      CONST_RETAIN_TIME_SNAP_SIGNAL : Time := t#200ms;   // Time retain snap signal to z300
      CONST_DWRIDPLATE : DWord := 16#20002;   // R_ID message
      CONST_DWRIDMESSAGE2 : DWord := 16#30003;   // R_ID message
      CONST_DWRIDMESSAGE : DWord := 16#10001;   // R_ID message
      CONST_DGLASSBREAK_CLASS : DInt := 5;   // Glass break used class
      CONST_DGLASSBREAK_SUBTYPE : DInt := 1002;   // Glass break subtype
      CONST_DGLASSBREAK_DEFECT_WIDTH_CMM : DInt := 366000;   // Defect width [mm/100]
      CONST_DGLASSBREAK_DEFECT_GAP_CMM : DInt := 40000;   // Glass break defect gap [mm/100]
      CONST_DGLASSBREAK_LASTDEFECT_LENGTH_CMM : DInt := 50000;   // Last defect on glass break length [mm/100]
   END_VAR
BEGIN

REGION Network 1: ####_CONSTANTS_####
END_REGION

REGION Network 2: ####_MATCH_####
END_REGION

REGION Network 3 (SCL): General reset clean
   IF #IN_xGeneralReset THEN

       #TMP_dwValue := 0;

       SCATTER(IN:=#TMP_dwValue,
               OUT=>#tPhases);

       SCATTER(IN:=#TMP_dwValue,
               OUT=>#tPhasesNetworkPlate);


   END_IF;
END_REGION

REGION Network 4 (SCL): Move data information to tracking
   #INO_tTrack.rgtTrackMachine[#IN_dMachineIndex].tUserData.dSetDistanceSnap_cmm := #IN_dSnapOffset_cmm*-1;
   #INO_tTrack.rgtTrackMachine[#IN_dMachineIndex].tUserData.dSetMachReacTime_ms := #tHMW.dAccelerationDelay_ms;
END_REGION

REGION Network 5 (SCL): Manage tracking call

   #OS_xNewCapUp := FALSE;
   #OS_xNewCapDw := FALSE;
   #OS_xNewCap := FALSE;
   #OS_xNewCapFastDropUp := FALSE;
   IF #INO_tTrack.rgtTrackMachine[#IN_dMachineIndex].tUserData.xGetPosReach THEN

       IF (NOT #ST_xPhaseInProgress) THEN

           IF #INO_tTrack.rgtTrackMachine[#IN_dMachineIndex].tUserData.dGetUpstremIndex >= 0 THEN
               #AUX_dUpCapIndex := #INO_tTrack.rgtTrackMachine[#IN_dMachineIndex].tUserData.dGetUpstremIndex;
               IF #INO_tTrack.rgtTrackCaps[#AUX_dUpCapIndex].tCap.dLength_cmm >= #CONST_MINPLATELENGTH_Z300_CMM THEN
                   #OS_xNewCapUp := TRUE;
                   #AUX_xValidUpCap := TRUE;
               ELSE
                   #AUX_xValidUpCap := FALSE;

               END_IF;
           ELSE
                   #AUX_xValidUpCap := FALSE;
                   #OS_xNewCapUp := FALSE;
                   #AUX_dUpCapIndex := 0;
           END_IF;

           IF #INO_tTrack.rgtTrackMachine[#IN_dMachineIndex].tUserData.dGetDownstreamIndex >= 0 THEN
               #AUX_xValidDwCap := TRUE;
               #OS_xNewCapDw := TRUE;            
               #AUX_dDwCapIndex := #INO_tTrack.rgtTrackMachine[#IN_dMachineIndex].tUserData.dGetDownstreamIndex;

               IF #INO_tTrack.rgtTrackCaps[#AUX_dDwCapIndex].tCap.dLength_cmm >= #CONST_MINPLATELENGTH_Z300_CMM THEN
                   #OS_xNewCap := TRUE;
               ELSE
                   #OS_xNewCapFastDropUp := TRUE;
               END_IF;

           ELSE
               #AUX_xValidDwCap := FALSE;
               #OS_xNewCapDw := FALSE;            
               #AUX_dDwCapIndex := 0;
           END_IF;



       END_IF;

       #INO_tTrack.rgtTrackMachine[#IN_dMachineIndex].tUserData.xGetPosReach := FALSE;

   END_IF;
END_REGION

REGION Network 6 (SCL): Manage message
   IF #AUX_xValidUpCap AND (#OS_xNewCapUp OR  #OS_xNewCapFastDropUp) THEN

       //Evaluate the missing xcut, send to cullet the upstream and downstream. On the downstream send also the message
       #TMP_xCutDone := FALSE;
       #AUX_xXcutDone := FALSE;
       FOR #TMP_dIndex := 0 TO "DMAXXHEADS_IND" DO
           IF #INO_tTrack.rgtTrackCaps[#AUX_dUpCapIndex].tCap.tDone.rgxXCutDoneHead[#TMP_dIndex] THEN
               #TMP_xCutDone := TRUE;
               #AUX_xXcutDone := TRUE;
               EXIT;                    
           END_IF;
       END_FOR;

       IF #TMP_xCutDone = FALSE THEN  

           //Send to cullet the upstream
           FOR #TMP_dIndex := 0 TO  #INO_tTrack.rgtTrackCaps[#AUX_dUpCapIndex].tCap.dNumLites - 1 DO

               IF #INO_tTrack.rgtTrackCaps[#AUX_dUpCapIndex].tCap.rgtLites[#TMP_dIndex].dMainDestination <> "DCULLETDESTMASK" THEN

                   #INO_tTrack.rgtTrackCaps[#AUX_dUpCapIndex].tCap.rgtLites[#TMP_dIndex].dMainDestination := "DCULLETDESTMASK";
                   #INO_tTrack.rgtTrackCaps[#AUX_dUpCapIndex].tCap.rgtLites[#TMP_dIndex].dAltDestination := 0;
                   #INO_tTrack.rgtTrackCaps[#AUX_dUpCapIndex].tCap.rgtLites[#TMP_dIndex].d2ndDestionation := 0;
                   #INO_tTrack.rgtTrackCaps[#AUX_dUpCapIndex].tCap.rgtLites[#TMP_dIndex].dCulletCause := "DCULLETCAUSE_XCUTMISSING";

               END_IF;
           END_FOR;

           #INO_tTrack.rgtTrackCaps[#AUX_dUpCapIndex].tCap.tRequests.xUpdateDataBPSA := TRUE;
           #INO_tTrack.rgtTrackCaps[#AUX_dUpCapIndex].tCap.tRequests.xUpdateDataBPSB := TRUE;

           //Send to cullet the downstream
           FOR #TMP_dIndex := 0 TO  #INO_tTrack.rgtTrackCaps[#AUX_dDwCapIndex].tCap.dNumLites - 1 DO

               IF #INO_tTrack.rgtTrackCaps[#AUX_dDwCapIndex].tCap.rgtLites[#TMP_dIndex].dMainDestination <> "DCULLETDESTMASK" THEN

                   #INO_tTrack.rgtTrackCaps[#AUX_dDwCapIndex].tCap.rgtLites[#TMP_dIndex].dMainDestination := "DCULLETDESTMASK";
                   #INO_tTrack.rgtTrackCaps[#AUX_dDwCapIndex].tCap.rgtLites[#TMP_dIndex].dAltDestination := 0;
                   #INO_tTrack.rgtTrackCaps[#AUX_dDwCapIndex].tCap.rgtLites[#TMP_dIndex].d2ndDestionation := 0;
                   #INO_tTrack.rgtTrackCaps[#AUX_dDwCapIndex].tCap.rgtLites[#TMP_dIndex].dCulletCause := "DCULLETCAUSE_XCUTMISSING";

                   "RP_AddMessageV2"(IN_xInit:=FALSE,
                     IN_dCodeEvent:="DEVENTS_REDESTINATION",
                     IN_strIndet_Max4Chars:='Z200',
                     IN_dValue1:="DEVENTS_CULLETDESTINATION",
                     IN_dValue2:=#INO_tTrack.rgtTrackCaps[#AUX_dDwCapIndex].tCap.rgtLites[#TMP_dIndex].dID,
                     IN_dValue3:=#INO_tTrack.rgtTrackCaps[#AUX_dDwCapIndex].tCap.rgtLites[#TMP_dIndex].dProductionID,
                     IN_dValue4:=#INO_tTrack.rgtTrackCaps[#AUX_dDwCapIndex].tCap.rgtLites[#TMP_dIndex].dCulletCause,
                     IN_dValue5:=0,
                     IN_dValue6:=0,
                     IN_dValue7:=0,
                     IN_dValue8:=0,
                     IN_dValue9:=0,
                     IN_dValue10:=0,
                     INO_tBuffer:=#INO_tMessage,
                     INO_xError:=#INO_xMessageAnomaly);

               END_IF;
           END_FOR;

           #INO_tTrack.rgtTrackCaps[#AUX_dUpCapIndex].tCap.tRequests.xUpdateDataBPSA := TRUE;
           #INO_tTrack.rgtTrackCaps[#AUX_dUpCapIndex].tCap.tRequests.xUpdateDataBPSB := TRUE;

       END_IF;

       FOR #TMP_dIndex := 0 TO #INO_tTrack.rgtTrackCaps[#AUX_dUpCapIndex].tCap.dNumLites - 1 DO

           IF #INO_tTrack.rgtTrackCaps[#AUX_dUpCapIndex].tCap.rgtLites[#TMP_dIndex].dMainDestination = "DCULLETDESTMASK" THEN
              "RP_AddMessageV2"(IN_xInit:=FALSE,
                     IN_dCodeEvent:="DEVENTS_REDESTINATION",
                     IN_strIndet_Max4Chars:='Z200',
                     IN_dValue1:="DEVENTS_CULLETDESTINATION",
                     IN_dValue2:=#INO_tTrack.rgtTrackCaps[#AUX_dUpCapIndex].tCap.rgtLites[#TMP_dIndex].dID,
                     IN_dValue3:=#INO_tTrack.rgtTrackCaps[#AUX_dUpCapIndex].tCap.rgtLites[#TMP_dIndex].dProductionID,
                     IN_dValue4:=#INO_tTrack.rgtTrackCaps[#AUX_dUpCapIndex].tCap.rgtLites[#TMP_dIndex].dCulletCause,
                     IN_dValue5:=0,
                     IN_dValue6:=0,
                     IN_dValue7:=0,
                     IN_dValue8:=0,
                     IN_dValue9:=0,
                     IN_dValue10:=0,
                     INO_tBuffer:=#INO_tMessage,
                     INO_xError:=#INO_xMessageAnomaly);
           END_IF;


       END_FOR;

   END_IF;
END_REGION

REGION Network 7: ####_HMI_LOGICS_####
END_REGION

REGION Network 8 (SCL): List of HMI logics
END_REGION

REGION Network 9: ####_ALARMS_####
END_REGION

REGION Network 10 (SCL): Reset alarms
   IF #IN_xResetAlarms THEN

       #TMP_dwValue := 0;

       SCATTER(IN:=#TMP_dwValue,
               OUT=>#tALM.tF);

       SCATTER(IN:=#TMP_dwValue,
               OUT=>#tALM.tS);

       SCATTER(IN:=#TMP_dwValue,
               OUT=>#tALM.tW);

   END_IF;
END_REGION

REGION Network 11: ####_STATUSES_####
END_REGION

REGION Network 12 (SCL): Calculate alarm statuses
   GATHER(IN:=#tALM.tS,
          OUT=>#TMP_dwValue);

   IF #TMP_dwValue <> 0 THEN
       #ST_xStoppingFaults := TRUE;
   ELSE
       #ST_xStoppingFaults := FALSE;
   END_IF;

   GATHER(IN:=#tALM.tF,
          OUT=>#TMP_dwValue);

   IF #TMP_dwValue <> 0 THEN
       #ST_xFaults := TRUE;
   ELSE
       #ST_xFaults := FALSE;
   END_IF;

   GATHER(IN:=#tALM.tW,
          OUT=>#TMP_dwValue);

   IF #TMP_dwValue <> 0 THEN
       #ST_xWarnings := TRUE;
   ELSE
       #ST_xWarnings := FALSE;
   END_IF;
END_REGION

REGION Network 13: Send data request
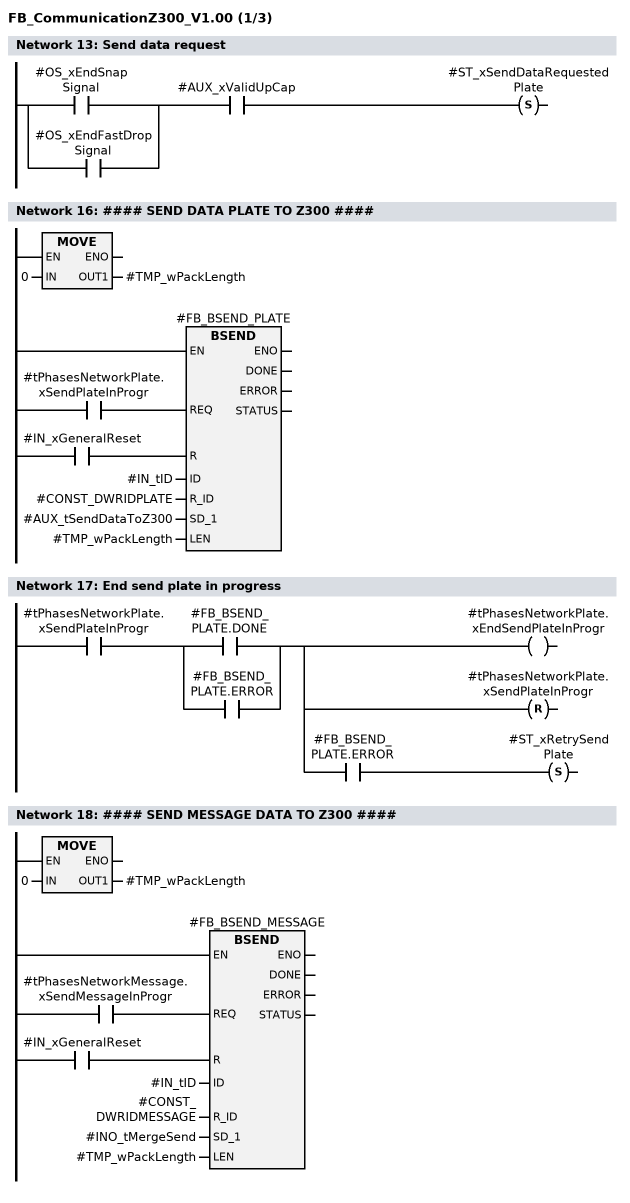
   RUNG wire#powerrail
      Contact( #OS_xEndSnapSignal )
      wire#w1
      Contact( #AUX_xValidUpCap )
      S_Coil( #ST_xSendDataRequestedPlate )
   END_RUNG
   RUNG wire#powerrail
      Contact( #OS_xEndFastDropSignal )
   END_RUNG wire#w1
   // the same network as SCL:
   IF (#OS_xEndSnapSignal OR #OS_xEndFastDropSignal) AND #AUX_xValidUpCap THEN
       #ST_xSendDataRequestedPlate := TRUE;
   END_IF;
END_REGION

REGION Network 14 (SCL): Compile Data for Z300
   IF NOT #ST_xPhaseInProgressNetworkPlate AND (#ST_xSendDataRequestedPlate OR #ST_xRetrySendPlate) THEN


       IF #ST_xSendDataRequestedPlate THEN

           //clean buffer
           #AUX_tSendDataToZ300 := #AUX_tEmptySendDataToZ300;
           //Convoy data.Search plate
           IF #INO_tTrack.rgtTrackCaps[#AUX_dUpCapIndex].tCap.dIndex = 0 THEN

               //Search until the previous cap
               #TMP_dIndex := 1;
               #TMP_dValue := #AUX_dUpCapIndex;
               #TMP_dConvNumPlate := 1;
               #TMP_dConvTotalLength_cmm := #INO_tTrack.rgtTrackCaps[#AUX_dUpCapIndex].tCap.dLength_cmm;

               WHILE #TMP_dIndex < "DMAXCAP_Z300" DO

                   #TMP_dValue := #TMP_dValue + 1;

                   IF #TMP_dValue > "DMAXTRACKCAP_IND" THEN
                       #TMP_dValue := 0;
                   END_IF;

                   IF #INO_tTrack.rgtTrackCaps[#TMP_dValue].tCap.dIndex <> 0 THEN

                       #TMP_dConvNumPlate := #TMP_dConvNumPlate + 1;
                       #TMP_dConvTotalLength_cmm := #TMP_dConvTotalLength_cmm + #INO_tTrack.rgtTrackCaps[#TMP_dValue].tCap.dLength_cmm;
                   ELSE

                       EXIT;

                   END_IF;

                   #TMP_dIndex := #TMP_dIndex + 1;

               END_WHILE;

               IF #TMP_dConvNumPlate > 1 THEN

                   //Convoy present, calculate gap.
                   #TMP_dConvGap_cmm := ("DMAXLENGHTCONVOY_CMM" - #TMP_dConvTotalLength_cmm) / (#TMP_dConvNumPlate - 1);
                   #TMP_dValue := #AUX_dUpCapIndex;
                   #TMP_dIndex := 0;
                   //Update plate data
                   WHILE (#TMP_dIndex < #TMP_dConvNumPlate) DO

                       #INO_tTrack.rgtTrackCaps[#TMP_dValue].tCap.dIndex := #TMP_dIndex;

                       IF (#TMP_dIndex + 1) < #TMP_dConvNumPlate THEN
                           #INO_tTrack.rgtTrackCaps[#TMP_dValue].tCap.dReqGapForConv_cmm := 50000; //#TMP_dConvGap_cmm;
                       ELSE
                           #INO_tTrack.rgtTrackCaps[#TMP_dValue].tCap.dReqGapForConv_cmm := 0;
                       END_IF;

                       #TMP_dIndex := #TMP_dIndex + 1;

                       #TMP_dValue := #TMP_dValue + 1;

                       IF #TMP_dValue > "DMAXTRACKCAP_IND"  THEN
                           #TMP_dValue := 0;
                       END_IF;

                   END_WHILE;
               END_IF;
           END_IF;

           #AUX_tCapToSend := #INO_tTrack.rgtTrackCaps[#AUX_dUpCapIndex].tCap;
           //compile plate data TO Z300
           #AUX_tSendDataToZ300.dID := #INO_tTrack.rgtTrackCaps[#AUX_dUpCapIndex].tCap.dID;
           #AUX_tSendDataToZ300.dProductionID := 1;
           #AUX_tSendDataToZ300.dLength_cmm := #INO_tTrack.rgtTrackCaps[#AUX_dUpCapIndex].tCap.dLength_cmm;
           #AUX_tSendDataToZ300.dWidth_cmm := #INO_tTrack.rgtTrackCaps[#AUX_dUpCapIndex].tCap.dWidth_cmm;
           #AUX_tSendDataToZ300.dThick_cmm := #INO_tTrack.rgtTrackCaps[#AUX_dUpCapIndex].tCap.dThick_cmm;
           #AUX_tSendDataToZ300.dIndex := #INO_tTrack.rgtTrackCaps[#AUX_dUpCapIndex].tCap.dIndex;
           #AUX_tSendDataToZ300.dFormat := #INO_tTrack.rgtTrackCaps[#AUX_dUpCapIndex].tCap.dFormat;
           #AUX_tSendDataToZ300.dNumLites := #INO_tTrack.rgtTrackCaps[#AUX_dUpCapIndex].tCap.dNumLites;

           #AUX_tSendDataToZ300.dReqGapForConv_cmm := 0;
           IF #INO_tTrack.rgtTrackCaps[#AUX_dUpCapIndex].tCap.dMaxCapInConv>1
               AND (#INO_tTrack.rgtTrackCaps[#AUX_dUpCapIndex].tCap.dMaxCapInConv-1>#AUX_tSendDataToZ300.dIndex) THEN
               #AUX_tSendDataToZ300.dReqGapForConv_cmm := 50000;
               #AUX_tSendDataToZ300.dGap_cmm := 50000;
           END_IF;
           #AUX_tSendDataToZ300.dMaxCapInConv := #INO_tTrack.rgtTrackCaps[#AUX_dUpCapIndex].tCap.dMaxCapInConv;

           #TMP_dValue := #AUX_dUpCapIndex + 1;

           IF #TMP_dValue >= "DMAXTRACKCAP_IND" THEN
               #TMP_dValue := 0;
           END_IF;
           IF #INO_tTrack.rgtTrackCaps[#TMP_dValue].tCap.dMaxCapInConv = 0 THEN
               #AUX_tSendDataToZ300.dReqGapForConv_cmm := 0;
               #AUX_tSendDataToZ300.dGap_cmm := 0;
               #AUX_tSendDataToZ300.dMaxCapInConv := 0;
           END_IF;


           #AUX_tSendDataToZ300.dConvTotLength_cmm := #INO_tTrack.rgtTrackCaps[#AUX_dUpCapIndex].tCap.dConvTotLength_cmm;
           #AUX_tSendDataToZ300.dMinWidth_cmm := #INO_tTrack.rgtTrackCaps[#AUX_dUpCapIndex].tCap.dMinWidth_cmm;
           #AUX_tSendDataToZ300.dMaxWidth_cmm := #INO_tTrack.rgtTrackCaps[#AUX_dUpCapIndex].tCap.dMaxWidth_cmm;
           #AUX_tSendDataToZ300.dGrossWidth_cmm := #INO_tTrack.rgtTrackCaps[#AUX_dUpCapIndex].tCap.dGrossWidth_cmm;
           #AUX_tSendDataToZ300.dNetWidth_cmm := #INO_tTrack.rgtTrackCaps[#AUX_dUpCapIndex].tCap.dNetWidth_cmm;
           #AUX_tSendDataToZ300.dDEdgeOpSide_cmm := #INO_tTrack.rgtTrackCaps[#AUX_dUpCapIndex].tCap.dDEdgeOpSide_cmm;
           #AUX_tSendDataToZ300.dDEdgeOppOpSide_cmm := #INO_tTrack.rgtTrackCaps[#AUX_dUpCapIndex].tCap.dDEdgeOppOpSide_cmm;
           #AUX_tSendDataToZ300.dTEdgeOpSide_cmm := #INO_tTrack.rgtTrackCaps[#AUX_dUpCapIndex].tCap.dTEdgeOpSide_cmm;
           #AUX_tSendDataToZ300.dTEdgeOppOpSide_cmm := #INO_tTrack.rgtTrackCaps[#AUX_dUpCapIndex].tCap.dTEdgeOppOpSide_cmm;
           #AUX_tSendDataToZ300.dCutWander_cmm := #INO_tTrack.rgtTrackCaps[#AUX_dUpCapIndex].tCap.dEndCutWander_cmm;
           #AUX_tSendDataToZ300.dColor := #INO_tTrack.rgtTrackCaps[#AUX_dUpCapIndex].tCap.dColor;
           #AUX_tSendDataToZ300.strColorDescr := #INO_tTrack.rgtTrackCaps[#AUX_dUpCapIndex].tCap.strColorDescr;

           #TMP_xReqDoneMatch := FALSE;
           GATHER(IN :=  #INO_tTrack.rgtTrackCaps[#AUX_dUpCapIndex].tCap.tDone.tYCuts[0].rgxHeadsDone,
                  OUT => #TMP_wValue);
           IF #TMP_wValue <> 0 THEN
               #AUX_tSendDataToZ300.tFlagTrim.xByYCut1 := TRUE;

               IF #INO_tTrack.rgtTrackCaps[#AUX_dUpCapIndex].tCap.tDone.tYCuts[0].rgxHeadsDone = 
                       #INO_tTrack.rgtTrackCaps[#AUX_dUpCapIndex].tCap.tRequests.tYCutsData[0].rgxHeadsRequest THEN
                   #TMP_xReqDoneMatch := TRUE;
               END_IF;

           END_IF;
           GATHER(IN := #INO_tTrack.rgtTrackCaps[#AUX_dUpCapIndex].tCap.tDone.tYCuts[1].rgxHeadsDone,
                  OUT => #TMP_wValue);
           IF #TMP_wValue <> 0 THEN
               #AUX_tSendDataToZ300.tFlagTrim.xByYCut2 := TRUE;

               IF #INO_tTrack.rgtTrackCaps[#AUX_dUpCapIndex].tCap.tDone.tYCuts[1].rgxHeadsDone = 
                       #INO_tTrack.rgtTrackCaps[#AUX_dUpCapIndex].tCap.tRequests.tYCutsData[1].rgxHeadsRequest THEN
                   #TMP_xReqDoneMatch := TRUE;
               END_IF;

           END_IF;

           IF #TMP_xReqDoneMatch THEN

               IF #INO_tTrack.rgtTrackCaps[#AUX_dUpCapIndex].tCap.dTEdgeOpSide_cmm > 0 THEN
                   #AUX_tSendDataToZ300.tFlagTrim.xTrim3OpSide := 1;
               END_IF;
               IF #INO_tTrack.rgtTrackCaps[#AUX_dUpCapIndex].tCap.dDEdgeOpSide_cmm > 0 THEN
                   #AUX_tSendDataToZ300.tFlagTrim.xTrim2OpSide := 1;
               END_IF;

               #AUX_tSendDataToZ300.tFlagTrim.xTrim1OpSide := 1;
               #AUX_tSendDataToZ300.tFlagTrim.xTrim1OppOpSide := 1;

               IF #INO_tTrack.rgtTrackCaps[#AUX_dUpCapIndex].tCap.dDEdgeOppOpSide_cmm > 0 THEN
                   #AUX_tSendDataToZ300.tFlagTrim.xTrim2OppOpSide := 1;
               END_IF;
               IF #INO_tTrack.rgtTrackCaps[#AUX_dUpCapIndex].tCap.dTEdgeOppOpSide_cmm > 0 THEN
                   #AUX_tSendDataToZ300.tFlagTrim.xTrim3OppOpSide := 1;
               END_IF;

               FOR #TMP_dIndex := 1 TO #INO_tTrack.rgtTrackCaps[#AUX_dUpCapIndex].tCap.dNumLites - 1 DO
                   #AUX_tSendDataToZ300.tFlagTrim.rgxIntCut[#TMP_dIndex - 1] := 1;
               END_FOR;

           ELSE
               #AUX_tSendDataToZ300.tFlagTrim.xTrim3OpSide := 0;
               #AUX_tSendDataToZ300.tFlagTrim.xTrim2OpSide := 0;
               #AUX_tSendDataToZ300.tFlagTrim.xTrim1OpSide := 0;
               #AUX_tSendDataToZ300.tFlagTrim.xTrim1OppOpSide := 0;
               #AUX_tSendDataToZ300.tFlagTrim.xTrim2OppOpSide := 0;
               #AUX_tSendDataToZ300.tFlagTrim.xTrim3OppOpSide := 0;
           END_IF;

           #AUX_tSendDataToZ300.tFlagTrim.xOptSelvedgeSel := #INO_tTrack.rgtTrackCaps[#AUX_dUpCapIndex].tCap.tRequests.xOptSelvedgeSel;
           #AUX_tSendDataToZ300.tFlagTrim.xOptSplitBarSel := #INO_tTrack.rgtTrackCaps[#AUX_dUpCapIndex].tCap.tRequests.xOptSplitBarSel;
           #AUX_tSendDataToZ300.tFlagTrim.xOptSepRollSel := #INO_tTrack.rgtTrackCaps[#AUX_dUpCapIndex].tCap.tRequests.xOptSepRollSel;

           FOR #TMP_dIndex := 0 TO "DMAXXHEADS_IND" DO
               #AUX_tSendDataToZ300.tFlagTrim.rgxXCutDoneHead[#TMP_dIndex] := #INO_tTrack.rgtTrackCaps[#AUX_dUpCapIndex].tCap.tDone.rgxXCutDoneHead[#TMP_dIndex];
           END_FOR;

           FOR #TMP_dIndex := 0 TO "DMAXXHEADS_IND" DO
               #AUX_tSendDataToZ300.tFlagTrim.rgxXCutDoneTail[#TMP_dIndex] := #INO_tTrack.rgtTrackCaps[#AUX_dUpCapIndex].tCap.tDone.rgxXCutDoneTail[#TMP_dIndex];
           END_FOR;

           IF #AUX_tSendDataToZ300.tFlagTrim.xByYCut1 THEN
               #AUX_tSendDataToZ300.tFlagTrim.rgxYCutHeadDone := #INO_tTrack.rgtTrackCaps[#AUX_dUpCapIndex].tCap.tDone.tYCuts[0].rgxHeadsDone;
           ELSE
               #AUX_tSendDataToZ300.tFlagTrim.rgxYCutHeadDone := #INO_tTrack.rgtTrackCaps[#AUX_dUpCapIndex].tCap.tDone.tYCuts[1].rgxHeadsDone;
           END_IF;

           #AUX_tSendDataToZ300.tFlagTrim.tSelvedge.dRequestTrim3OpSide := #INO_tTrack.rgtTrackCaps[#AUX_dUpCapIndex].tCap.tRequests.dReqTrim3OpSide;
           #AUX_tSendDataToZ300.tFlagTrim.tSelvedge.dRequestTrim2OpSide := #INO_tTrack.rgtTrackCaps[#AUX_dUpCapIndex].tCap.tRequests.dReqTrim2OpSide;
           #AUX_tSendDataToZ300.tFlagTrim.tSelvedge.dRequestTrim1OpSide := #INO_tTrack.rgtTrackCaps[#AUX_dUpCapIndex].tCap.tRequests.dReqTrim1OpSide;
           #AUX_tSendDataToZ300.tFlagTrim.tSelvedge.dRequestTrim3OppOpSide := #INO_tTrack.rgtTrackCaps[#AUX_dUpCapIndex].tCap.tRequests.dReqTrim3OppOpSide;
           #AUX_tSendDataToZ300.tFlagTrim.tSelvedge.dRequestTrim2OppOpSide := #INO_tTrack.rgtTrackCaps[#AUX_dUpCapIndex].tCap.tRequests.dReqTrim2OppOpSide;
           #AUX_tSendDataToZ300.tFlagTrim.tSelvedge.dRequestTrim1OppOpSide := #INO_tTrack.rgtTrackCaps[#AUX_dUpCapIndex].tCap.tRequests.dReqTrim1OppOpSide;

           FOR #TMP_dIndex := 0 TO "DMAXLITE_IND" DO
               #AUX_tSendDataToZ300.tFlagTrim.tSplitBar[#TMP_dIndex].dRequestSnapCut := #INO_tTrack.rgtTrackCaps[#AUX_dUpCapIndex].tCap.tRequests.rgdReqSplitBarSel[#TMP_dIndex];
           END_FOR;

           FOR #TMP_dIndex := 0 TO "DMAXSEPROLLBANK_IND" DO
               #TMP_wValue := INT_TO_WORD(#INO_tTrack.rgtTrackCaps[#AUX_dUpCapIndex].tCap.tRequests.rgbSeparatorSelect[#TMP_dIndex]);
               SCATTER(IN := #TMP_wValue,
                       OUT => #TMP_rgxWValue);
               #AUX_tSendDataToZ300.tFlagTrim.tSepRoll[#TMP_dIndex].rgxRequestSeparator := #TMP_rgxWValue;
           END_FOR;

           FOR #TMP_dIndex := 0 TO "DMAXLITE_Z300"  DO
               #AUX_tSendDataToZ300.rgtLites[#TMP_dIndex].dID := #INO_tTrack.rgtTrackCaps[#AUX_dUpCapIndex].tCap.rgtLites[#TMP_dIndex].dID;
               #AUX_tSendDataToZ300.rgtLites[#TMP_dIndex].dProductionID := #INO_tTrack.rgtTrackCaps[#AUX_dUpCapIndex].tCap.rgtLites[#TMP_dIndex].dProductionID;
               #AUX_tSendDataToZ300.rgtLites[#TMP_dIndex].strProdDescr := #INO_tTrack.rgtTrackCaps[#AUX_dUpCapIndex].tCap.rgtLites[#TMP_dIndex].strProdDescr;
               #AUX_tSendDataToZ300.rgtLites[#TMP_dIndex].dQualityID := #INO_tTrack.rgtTrackCaps[#AUX_dUpCapIndex].tCap.rgtLites[#TMP_dIndex].dQualityID;
               #AUX_tSendDataToZ300.rgtLites[#TMP_dIndex].strQualityDescr := #INO_tTrack.rgtTrackCaps[#AUX_dUpCapIndex].tCap.rgtLites[#TMP_dIndex].strQualityDescr;
               #AUX_tSendDataToZ300.rgtLites[#TMP_dIndex].dCameraRecipeID := #INO_tTrack.rgtTrackCaps[#AUX_dUpCapIndex].tCap.rgtLites[#TMP_dIndex].dCameraRecipeID;
               #AUX_tSendDataToZ300.rgtLites[#TMP_dIndex].dWidth_cmm := #INO_tTrack.rgtTrackCaps[#AUX_dUpCapIndex].tCap.rgtLites[#TMP_dIndex].dWidth_cmm;
               #AUX_tSendDataToZ300.rgtLites[#TMP_dIndex].dBarycentre_cmm := #INO_tTrack.rgtTrackCaps[#AUX_dUpCapIndex].tCap.rgtLites[#TMP_dIndex].dBarycentre_cmm ;
               #AUX_tSendDataToZ300.rgtLites[#TMP_dIndex].dCulletCause_cmm := #INO_tTrack.rgtTrackCaps[#AUX_dUpCapIndex].tCap.rgtLites[#TMP_dIndex].dCulletCause;
               #AUX_tSendDataToZ300.rgtLites[#TMP_dIndex].tRequests.xReqGeoIspection := #INO_tTrack.rgtTrackCaps[#AUX_dUpCapIndex].tCap.rgtLites[#TMP_dIndex].tRequests.xGeomInsp;
               #AUX_tSendDataToZ300.rgtLites[#TMP_dIndex].tRequests.xReqPowderA := #INO_tTrack.rgtTrackCaps[#AUX_dUpCapIndex].tCap.rgtLites[#TMP_dIndex].rgxLayers[0];
               #AUX_tSendDataToZ300.rgtLites[#TMP_dIndex].tRequests.xReqPowderB := #INO_tTrack.rgtTrackCaps[#AUX_dUpCapIndex].tCap.rgtLites[#TMP_dIndex].rgxLayers[1];
               #AUX_tSendDataToZ300.rgtLites[#TMP_dIndex].tRequests.Spare4 := #INO_tTrack.rgtTrackCaps[#AUX_dUpCapIndex].tCap.rgtLites[#TMP_dIndex].rgxLayers[0];
               #AUX_tSendDataToZ300.rgtLites[#TMP_dIndex].xSaturationPlate := #INO_tTrack.rgtTrackCaps[#AUX_dUpCapIndex].tCap.rgtLites[#TMP_dIndex].xSaturationPlate;

               #TMP_lwValue := LINT_TO_LWORD(#INO_tTrack.rgtTrackCaps[#AUX_dUpCapIndex].tCap.rgtLites[#TMP_dIndex].dMainDestination);
               SCATTER(IN := #TMP_lwValue,
                       OUT => #AUX_tSendDataToZ300.rgtLites[#TMP_dIndex].rgxMain);

               #TMP_lwValue := LINT_TO_LWORD(#INO_tTrack.rgtTrackCaps[#AUX_dUpCapIndex].tCap.rgtLites[#TMP_dIndex].dAltDestination);
               SCATTER(IN := #TMP_lwValue,
                       OUT => #AUX_tSendDataToZ300.rgtLites[#TMP_dIndex].rgxAlternative);


               #TMP_lwValue := LINT_TO_LWORD(#INO_tTrack.rgtTrackCaps[#AUX_dUpCapIndex].tCap.rgtLites[#TMP_dIndex].d2ndDestionation);
               SCATTER(IN := #TMP_lwValue,
                       OUT => #AUX_tSendDataToZ300.rgtLites[#TMP_dIndex].rgx2ndDestination);


           END_FOR;

           #tPhasesNetworkPlate.xSendPlateInProgr := TRUE;
           #ST_xSendDataRequestedPlate := 0;
       END_IF;

       IF #ST_xRetrySendPlate = TRUE THEN
           #tPhasesNetworkPlate.xSendPlateInProgr := TRUE;
           #ST_xRetrySendPlate := FALSE;
       END_IF;

   END_IF;
END_REGION

REGION Network 15 (SCL): Check if a new message packet is request to send
   IF NOT #ST_xPhaseInProgressNetworkMessage AND #INO_tMergeSend.xInitialized AND #INO_tMergeSend.dNumOfMessage > 0 THEN

       #tPhasesNetworkMessage.xSendMessageInProgr := TRUE;

       //Analyze the message. If some change destinationation is required check if the plate is still on z200 buffer
       FOR #TMP_dMexIndex := 0 TO #INO_tMergeSend.dNumOfMessage - 1 DO
           #TMP_xExit := FALSE;
           IF (#INO_tMergeSend.rgtMessages[#TMP_dMexIndex].dCodeEvent = "DEVENTS_REDEST_OPT") THEN

               //Search the plate on buffer
               #TMP_dTrackTail := #INO_tTrack.dTrackingTail;

               WHILE (#TMP_dTrackTail <> #INO_tTrack.dTrackingHead) AND NOT #TMP_xExit DO

                   FOR #TMP_dIndex := 0 TO #INO_tTrack.rgtTrackCaps[#TMP_dTrackTail].tCap.dNumLites -1 DO

                       IF (#INO_tTrack.rgtTrackCaps[#TMP_dTrackTail].tCap.rgtLites[#TMP_dIndex].dID = #INO_tMergeSend.rgtMessages[#TMP_dMexIndex].dEvent1) THEN

                           #INO_tTrack.rgtTrackCaps[#TMP_dTrackTail].tCap.rgtLites[#TMP_dIndex].dMainDestination := 2 ** #INO_tMergeSend.rgtMessages[#TMP_dMexIndex].dEvent4;
                           #INO_tTrack.rgtTrackCaps[#TMP_dTrackTail].tCap.rgtLites[#TMP_dIndex].dCulletCause := #INO_tMergeSend.rgtMessages[#TMP_dMexIndex].dEvent3;
                           #INO_tTrack.rgtTrackCaps[#TMP_dTrackTail].tCap.tRequests.xUpdateDataBPSA := TRUE;
                           #INO_tTrack.rgtTrackCaps[#TMP_dTrackTail].tCap.tRequests.xUpdateDataBPSB := TRUE;
                           #TMP_xExit := TRUE;
                           EXIT;    
                       END_IF;  

                   END_FOR;

                   IF (#TMP_dTrackTail + 1) >= "DMAXTRACKCAP" THEN
                       #TMP_dTrackTail := 0;
                   ELSE
                       #TMP_dTrackTail += 1;
                   END_IF;

               END_WHILE;

           END_IF;

       END_FOR;
       //#INO_tMergeSend.dNumOfMessage := 0;

   END_IF;
END_REGION

REGION Network 16: #### SEND DATA PLATE TO Z300 ####
   #TMP_wPackLength := 0;
   #FB_BSEND_PLATE(REQ := #tPhasesNetworkPlate.xSendPlateInProgr,   // BSEND
                   R := #IN_xGeneralReset,
                   ID := #IN_tID,
                   R_ID := #CONST_DWRIDPLATE,
                   SD_1 := #AUX_tSendDataToZ300,
                   LEN := #TMP_wPackLength);
END_REGION

REGION Network 17: End send plate in progress
   RUNG wire#powerrail
      Contact( #tPhasesNetworkPlate.xSendPlateInProgr )
      wire#w1
      Contact( #FB_BSEND_PLATE.DONE )
      wire#w2
      Coil( #tPhasesNetworkPlate.xEndSendPlateInProgr )
   END_RUNG
   RUNG wire#w1
      Contact( #FB_BSEND_PLATE.ERROR )
   END_RUNG wire#w2
   RUNG wire#w2
      R_Coil( #tPhasesNetworkPlate.xSendPlateInProgr )
   END_RUNG
   RUNG wire#w2
      Contact( #FB_BSEND_PLATE.ERROR )
      S_Coil( #ST_xRetrySendPlate )
   END_RUNG
   // the same network as SCL:
   #tPhasesNetworkPlate.xEndSendPlateInProgr := #tPhasesNetworkPlate.xSendPlateInProgr AND (#FB_BSEND_PLATE.DONE OR #FB_BSEND_PLATE.ERROR);
   IF #tPhasesNetworkPlate.xEndSendPlateInProgr THEN #tPhasesNetworkPlate.xSendPlateInProgr := FALSE; END_IF;
   IF #tPhasesNetworkPlate.xEndSendPlateInProgr AND #FB_BSEND_PLATE.ERROR THEN
       #ST_xRetrySendPlate := TRUE;
   END_IF;
END_REGION

REGION Network 18: #### SEND MESSAGE DATA TO Z300 ####
   #TMP_wPackLength := 0;
   #FB_BSEND_MESSAGE(REQ := #tPhasesNetworkMessage.xSendMessageInProgr,   // BSEND
                     R := #IN_xGeneralReset,
                     ID := #IN_tID,
                     R_ID := #CONST_DWRIDMESSAGE,
                     SD_1 := #INO_tMergeSend,
                     LEN := #TMP_wPackLength);
END_REGION

REGION Network 19: End send msg in progress
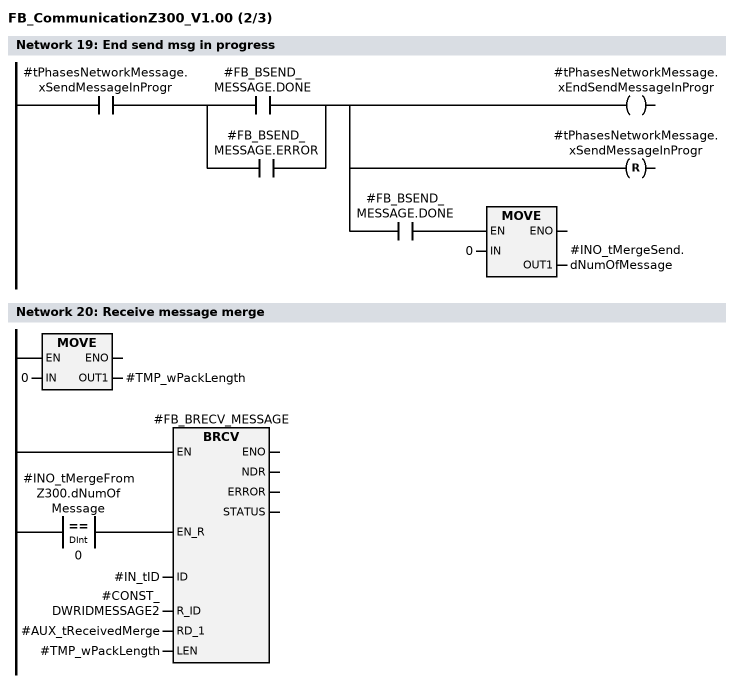
   RUNG wire#powerrail
      Contact( #tPhasesNetworkMessage.xSendMessageInProgr )
      wire#w1
      Contact( #FB_BSEND_MESSAGE.DONE )
      wire#w2
      Coil( #tPhasesNetworkMessage.xEndSendMessageInProgr )
   END_RUNG
   RUNG wire#w1
      Contact( #FB_BSEND_MESSAGE.ERROR )
   END_RUNG wire#w2
   RUNG wire#w2
      R_Coil( #tPhasesNetworkMessage.xSendMessageInProgr )
   END_RUNG
   RUNG wire#w2
      Contact( #FB_BSEND_MESSAGE.DONE )
      Move(in := 0, out1 => #INO_tMergeSend.dNumOfMessage)
   END_RUNG
   // the same network as SCL:
   #tPhasesNetworkMessage.xEndSendMessageInProgr := #tPhasesNetworkMessage.xSendMessageInProgr AND (#FB_BSEND_MESSAGE.DONE OR #FB_BSEND_MESSAGE.ERROR);
   IF #tPhasesNetworkMessage.xEndSendMessageInProgr THEN
       #tPhasesNetworkMessage.xSendMessageInProgr := FALSE;
   END_IF;
   IF #tPhasesNetworkMessage.xEndSendMessageInProgr AND #FB_BSEND_MESSAGE.DONE THEN
       #INO_tMergeSend.dNumOfMessage := 0;
   END_IF;
END_REGION

REGION Network 20: Receive message merge
   #TMP_wPackLength := 0;
   #FB_BRECV_MESSAGE(EN_R := #INO_tMergeFromZ300.dNumOfMessage = 0,   // BRCV
                     ID := #IN_tID,
                     R_ID := #CONST_DWRIDMESSAGE2,
                     RD_1 := #AUX_tReceivedMerge,
                     LEN := #TMP_wPackLength);
END_REGION

REGION Network 21 (SCL): Manage received data
   IF #FB_BRECV_MESSAGE.NDR THEN

       IF #AUX_tReceivedMerge.dNumOfMessage > 0 THEN

           #TMP_dNumMessage := #AUX_tReceivedMerge.dNumOfMessage;
           #INO_tMergeFromZ300 := #AUX_tReceivedMerge;
           #INO_tMergeFromZ300.dNumOfMessage := #TMP_dNumMessage;
       END_IF;

   END_IF;
END_REGION

REGION Network 22 (SCL): Calculare phase in progress
   GATHER(IN:=#tPhases,
          OUT=>#TMP_dwValue);

   IF #TMP_dwValue <> 0 THEN
       #ST_xPhaseInProgress := TRUE;
   ELSE
       #ST_xPhaseInProgress := FALSE;
   END_IF;

   GATHER(IN := #tPhasesNetworkPlate,
           OUT => #TMP_dwValue);

   IF  #TMP_dwValue <> 0 THEN
       #ST_xPhaseInProgressNetworkPlate := TRUE;
   ELSE
       #ST_xPhaseInProgressNetworkPlate := FALSE;
   END_IF;

   GATHER(IN := #tPhasesNetworkMessage,
           OUT => #TMP_dwValue);

   IF #TMP_dwValue <> 0 THEN
       #ST_xPhaseInProgressNetworkMessage := TRUE;
   ELSE
       #ST_xPhaseInProgressNetworkMessage := FALSE;
   END_IF;
END_REGION

REGION Network 23: ####_OUTPUT_####
END_REGION

REGION Network 24: Idevice outputs
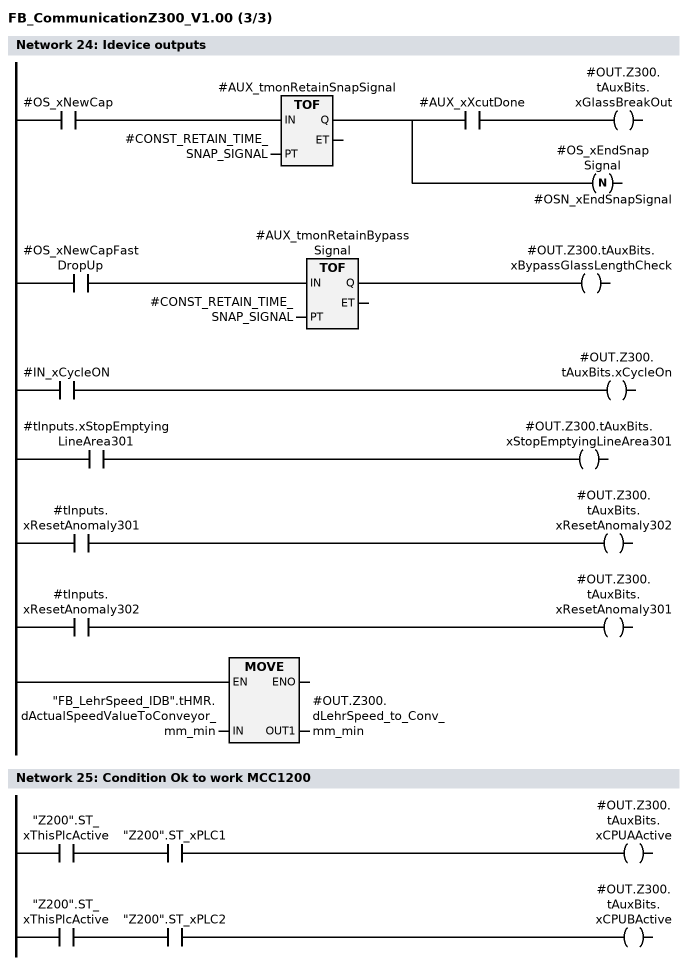
   #AUX_tmonRetainSnapSignal(IN := #OS_xNewCap, PT := #CONST_RETAIN_TIME_SNAP_SIGNAL);   // TOF
   #OUT.Z300.tAuxBits.xGlassBreakOut := #AUX_tmonRetainSnapSignal.Q AND #AUX_xXcutDone;
   #OS_xEndSnapSignal := NOT #AUX_tmonRetainSnapSignal.Q AND #OSN_xEndSnapSignal;   // falling edge
   #OSN_xEndSnapSignal := #AUX_tmonRetainSnapSignal.Q;
   #AUX_tmonRetainBypassSignal(IN := #OS_xNewCapFastDropUp, PT := #CONST_RETAIN_TIME_SNAP_SIGNAL);   // TOF
   #OUT.Z300.tAuxBits.xBypassGlassLengthCheck := #AUX_tmonRetainBypassSignal.Q;
   #OUT.Z300.tAuxBits.xCycleOn := #IN_xCycleON;
   #OUT.Z300.tAuxBits.xStopEmptyingLineArea301 := #tInputs.xStopEmptyingLineArea301;
   #OUT.Z300.tAuxBits.xResetAnomaly302 := #tInputs.xResetAnomaly301;
   #OUT.Z300.tAuxBits.xResetAnomaly301 := #tInputs.xResetAnomaly302;
   #OUT.Z300.dLehrSpeed_to_Conv_mm_min := "FB_LehrSpeed_IDB".tHMR.dActualSpeedValueToConveyor_mm_min;
END_REGION

REGION Network 25: Condition Ok to work MCC1200
   RUNG wire#powerrail
      Contact( "Z200".ST_xThisPlcActive )
      Contact( "Z200".ST_xPLC1 )
      Coil( #OUT.Z300.tAuxBits.xCPUAActive )
   END_RUNG
   RUNG wire#powerrail
      Contact( "Z200".ST_xThisPlcActive )
      Contact( "Z200".ST_xPLC2 )
      Coil( #OUT.Z300.tAuxBits.xCPUBActive )
   END_RUNG
   // the same network as SCL:
   #OUT.Z300.tAuxBits.xCPUAActive := "Z200".ST_xThisPlcActive AND "Z200".ST_xPLC1;
   #OUT.Z300.tAuxBits.xCPUBActive := "Z200".ST_xThisPlcActive AND "Z200".ST_xPLC2;
END_REGION
END_FUNCTION_BLOCK

// folder: 03_Programs_Logics/MCC1200/14_BPS

